// TIA Portal project "SSA-3GHz_V18" (V18) (continued)
REGION Network 4: INFO: If T_CONFIG is done, "start" will be reset.
   RUNG wire#powerrail
      { S7_Templates := "SrcType := DWord" } EQ_Contact(in1 := "SLI_gDB_T_CONFIG_PLC".T_CONFIG.status, in2 := 16#0070_0200)
      R_Coil( "SLI_gDB_T_CONFIG_PLC".T_CONFIG.start )
   END_RUNG
   // the same network as SCL:
   IF "SLI_gDB_T_CONFIG_PLC".T_CONFIG.status = 16#0070_0200 THEN
       "SLI_gDB_T_CONFIG_PLC".T_CONFIG.start := FALSE;
   END_IF;
END_REGION
END_FUNCTION

FUNCTION "ProcessDI" : Void   // FC400, LAD
{ S7_Optimized_Access := 'TRUE' }
VERSION : 0.1
BEGIN

REGION Network 1: DutyCycOK
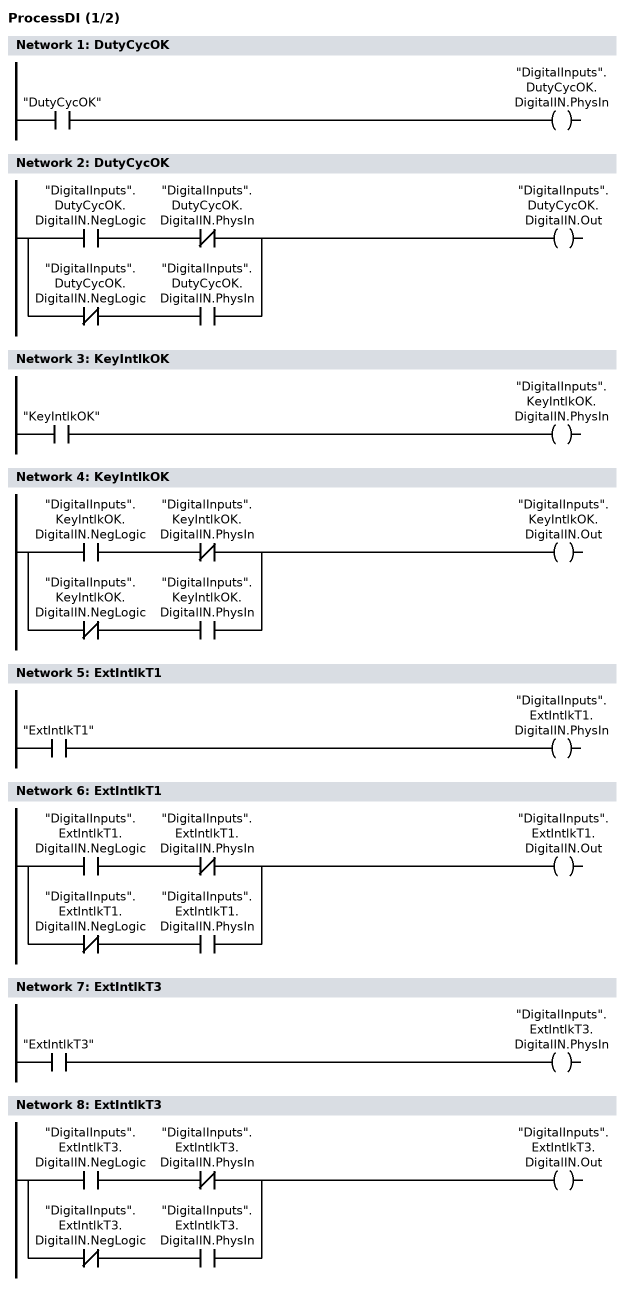
   RUNG wire#powerrail
      Contact( "DutyCycOK" )
      Coil( "DigitalInputs".DutyCycOK.DigitalIN.PhysIn )
   END_RUNG
   // the same network as SCL:
   "DigitalInputs".DutyCycOK.DigitalIN.PhysIn := "DutyCycOK";
END_REGION

REGION Network 2: DutyCycOK
   RUNG wire#powerrail
      Contact( "DigitalInputs".DutyCycOK.DigitalIN.NegLogic )
      I_Contact( "DigitalInputs".DutyCycOK.DigitalIN.PhysIn )
      wire#w1
      Coil( "DigitalInputs".DutyCycOK.DigitalIN.Out )
   END_RUNG
   RUNG wire#powerrail
      I_Contact( "DigitalInputs".DutyCycOK.DigitalIN.NegLogic )
      Contact( "DigitalInputs".DutyCycOK.DigitalIN.PhysIn )
   END_RUNG wire#w1
   // the same network as SCL:
   "DigitalInputs".DutyCycOK.DigitalIN.Out := ("DigitalInputs".DutyCycOK.DigitalIN.NegLogic AND NOT "DigitalInputs".DutyCycOK.DigitalIN.PhysIn) OR (NOT "DigitalInputs".DutyCycOK.DigitalIN.NegLogic AND "DigitalInputs".DutyCycOK.DigitalIN.PhysIn);
END_REGION

REGION Network 3: KeyIntlkOK
   RUNG wire#powerrail
      Contact( "KeyIntlkOK" )
      Coil( "DigitalInputs".KeyIntlkOK.DigitalIN.PhysIn )
   END_RUNG
   // the same network as SCL:
   "DigitalInputs".KeyIntlkOK.DigitalIN.PhysIn := "KeyIntlkOK";
END_REGION

REGION Network 4: KeyIntlkOK
   RUNG wire#powerrail
      Contact( "DigitalInputs".KeyIntlkOK.DigitalIN.NegLogic )
      I_Contact( "DigitalInputs".KeyIntlkOK.DigitalIN.PhysIn )
      wire#w1
      Coil( "DigitalInputs".KeyIntlkOK.DigitalIN.Out )
   END_RUNG
   RUNG wire#powerrail
      I_Contact( "DigitalInputs".KeyIntlkOK.DigitalIN.NegLogic )
      Contact( "DigitalInputs".KeyIntlkOK.DigitalIN.PhysIn )
   END_RUNG wire#w1
   // the same network as SCL:
   "DigitalInputs".KeyIntlkOK.DigitalIN.Out := ("DigitalInputs".KeyIntlkOK.DigitalIN.NegLogic AND NOT "DigitalInputs".KeyIntlkOK.DigitalIN.PhysIn) OR (NOT "DigitalInputs".KeyIntlkOK.DigitalIN.NegLogic AND "DigitalInputs".KeyIntlkOK.DigitalIN.PhysIn);
END_REGION

REGION Network 5: ExtIntlkT1
   RUNG wire#powerrail
      Contact( "ExtIntlkT1" )
      Coil( "DigitalInputs".ExtIntlkT1.DigitalIN.PhysIn )
   END_RUNG
   // the same network as SCL:
   "DigitalInputs".ExtIntlkT1.DigitalIN.PhysIn := "ExtIntlkT1";
END_REGION

REGION Network 6: ExtIntlkT1
   RUNG wire#powerrail
      Contact( "DigitalInputs".ExtIntlkT1.DigitalIN.NegLogic )
      I_Contact( "DigitalInputs".ExtIntlkT1.DigitalIN.PhysIn )
      wire#w1
      Coil( "DigitalInputs".ExtIntlkT1.DigitalIN.Out )
   END_RUNG
   RUNG wire#powerrail
      I_Contact( "DigitalInputs".ExtIntlkT1.DigitalIN.NegLogic )
      Contact( "DigitalInputs".ExtIntlkT1.DigitalIN.PhysIn )
   END_RUNG wire#w1
   // the same network as SCL:
   "DigitalInputs".ExtIntlkT1.DigitalIN.Out := ("DigitalInputs".ExtIntlkT1.DigitalIN.NegLogic AND NOT "DigitalInputs".ExtIntlkT1.DigitalIN.PhysIn) OR (NOT "DigitalInputs".ExtIntlkT1.DigitalIN.NegLogic AND "DigitalInputs".ExtIntlkT1.DigitalIN.PhysIn);
END_REGION

REGION Network 7: ExtIntlkT3
   RUNG wire#powerrail
      Contact( "ExtIntlkT3" )
      Coil( "DigitalInputs".ExtIntlkT3.DigitalIN.PhysIn )
   END_RUNG
   // the same network as SCL:
   "DigitalInputs".ExtIntlkT3.DigitalIN.PhysIn := "ExtIntlkT3";
END_REGION

REGION Network 8: ExtIntlkT3
   RUNG wire#powerrail
      Contact( "DigitalInputs".ExtIntlkT3.DigitalIN.NegLogic )
      I_Contact( "DigitalInputs".ExtIntlkT3.DigitalIN.PhysIn )
      wire#w1
      Coil( "DigitalInputs".ExtIntlkT3.DigitalIN.Out )
   END_RUNG
   RUNG wire#powerrail
      I_Contact( "DigitalInputs".ExtIntlkT3.DigitalIN.NegLogic )
      Contact( "DigitalInputs".ExtIntlkT3.DigitalIN.PhysIn )
   END_RUNG wire#w1
   // the same network as SCL:
   "DigitalInputs".ExtIntlkT3.DigitalIN.Out := ("DigitalInputs".ExtIntlkT3.DigitalIN.NegLogic AND NOT "DigitalInputs".ExtIntlkT3.DigitalIN.PhysIn) OR (NOT "DigitalInputs".ExtIntlkT3.DigitalIN.NegLogic AND "DigitalInputs".ExtIntlkT3.DigitalIN.PhysIn);
END_REGION

REGION Network 9: PS_OK
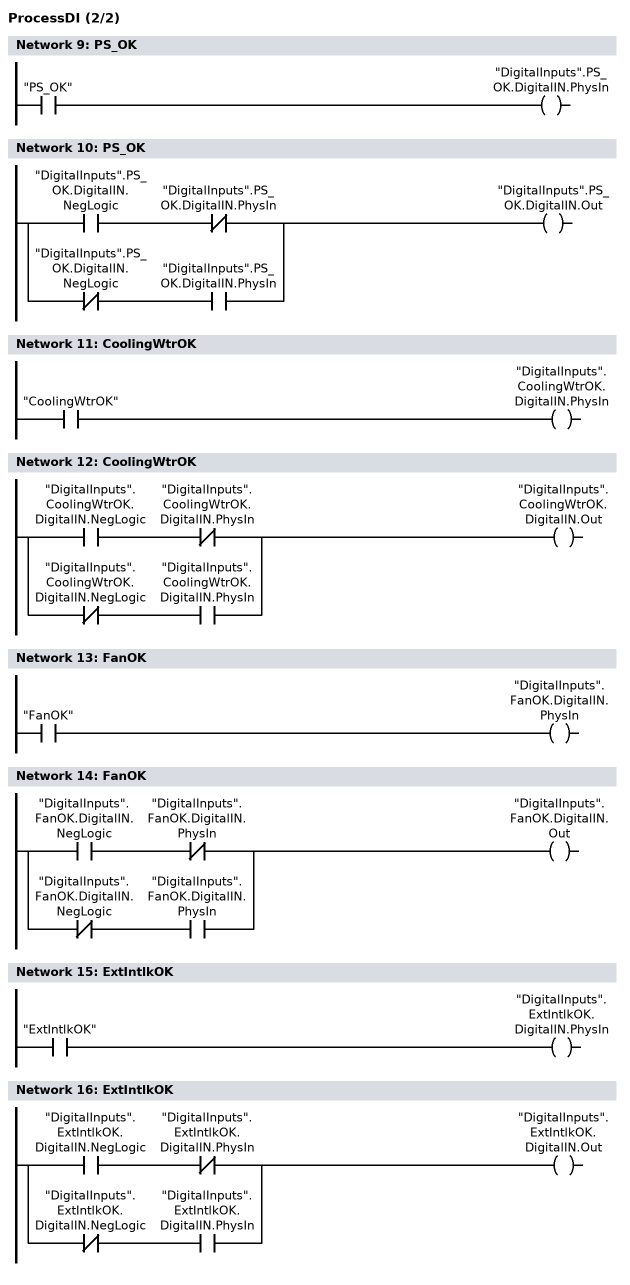
   RUNG wire#powerrail
      Contact( "PS_OK" )
      Coil( "DigitalInputs".PS_OK.DigitalIN.PhysIn )
   END_RUNG
   // the same network as SCL:
   "DigitalInputs".PS_OK.DigitalIN.PhysIn := "PS_OK";
END_REGION

REGION Network 10: PS_OK
   RUNG wire#powerrail
      Contact( "DigitalInputs".PS_OK.DigitalIN.NegLogic )
      I_Contact( "DigitalInputs".PS_OK.DigitalIN.PhysIn )
      wire#w1
      Coil( "DigitalInputs".PS_OK.DigitalIN.Out )
   END_RUNG
   RUNG wire#powerrail
      I_Contact( "DigitalInputs".PS_OK.DigitalIN.NegLogic )
      Contact( "DigitalInputs".PS_OK.DigitalIN.PhysIn )
   END_RUNG wire#w1
   // the same network as SCL:
   "DigitalInputs".PS_OK.DigitalIN.Out := ("DigitalInputs".PS_OK.DigitalIN.NegLogic AND NOT "DigitalInputs".PS_OK.DigitalIN.PhysIn) OR (NOT "DigitalInputs".PS_OK.DigitalIN.NegLogic AND "DigitalInputs".PS_OK.DigitalIN.PhysIn);
END_REGION

REGION Network 11: CoolingWtrOK
   RUNG wire#powerrail
      Contact( "CoolingWtrOK" )
      Coil( "DigitalInputs".CoolingWtrOK.DigitalIN.PhysIn )
   END_RUNG
   // the same network as SCL:
   "DigitalInputs".CoolingWtrOK.DigitalIN.PhysIn := "CoolingWtrOK";
END_REGION

REGION Network 12: CoolingWtrOK
   RUNG wire#powerrail
      Contact( "DigitalInputs".CoolingWtrOK.DigitalIN.NegLogic )
      I_Contact( "DigitalInputs".CoolingWtrOK.DigitalIN.PhysIn )
      wire#w1
      Coil( "DigitalInputs".CoolingWtrOK.DigitalIN.Out )
   END_RUNG
   RUNG wire#powerrail
      I_Contact( "DigitalInputs".CoolingWtrOK.DigitalIN.NegLogic )
      Contact( "DigitalInputs".CoolingWtrOK.DigitalIN.PhysIn )
   END_RUNG wire#w1
   // the same network as SCL:
   "DigitalInputs".CoolingWtrOK.DigitalIN.Out := ("DigitalInputs".CoolingWtrOK.DigitalIN.NegLogic AND NOT "DigitalInputs".CoolingWtrOK.DigitalIN.PhysIn) OR (NOT "DigitalInputs".CoolingWtrOK.DigitalIN.NegLogic AND "DigitalInputs".CoolingWtrOK.DigitalIN.PhysIn);
END_REGION

REGION Network 13: FanOK
   RUNG wire#powerrail
      Contact( "FanOK" )
      Coil( "DigitalInputs".FanOK.DigitalIN.PhysIn )
   END_RUNG
   // the same network as SCL:
   "DigitalInputs".FanOK.DigitalIN.PhysIn := "FanOK";
END_REGION

REGION Network 14: FanOK
   RUNG wire#powerrail
      Contact( "DigitalInputs".FanOK.DigitalIN.NegLogic )
      I_Contact( "DigitalInputs".FanOK.DigitalIN.PhysIn )
      wire#w1
      Coil( "DigitalInputs".FanOK.DigitalIN.Out )
   END_RUNG
   RUNG wire#powerrail
      I_Contact( "DigitalInputs".FanOK.DigitalIN.NegLogic )
      Contact( "DigitalInputs".FanOK.DigitalIN.PhysIn )
   END_RUNG wire#w1
   // the same network as SCL:
   "DigitalInputs".FanOK.DigitalIN.Out := ("DigitalInputs".FanOK.DigitalIN.NegLogic AND NOT "DigitalInputs".FanOK.DigitalIN.PhysIn) OR (NOT "DigitalInputs".FanOK.DigitalIN.NegLogic AND "DigitalInputs".FanOK.DigitalIN.PhysIn);
END_REGION

REGION Network 15: ExtIntlkOK
   RUNG wire#powerrail
      Contact( "ExtIntlkOK" )
      Coil( "DigitalInputs".ExtIntlkOK.DigitalIN.PhysIn )
   END_RUNG
   // the same network as SCL:
   "DigitalInputs".ExtIntlkOK.DigitalIN.PhysIn := "ExtIntlkOK";
END_REGION

REGION Network 16: ExtIntlkOK
   RUNG wire#powerrail
      Contact( "DigitalInputs".ExtIntlkOK.DigitalIN.NegLogic )
      I_Contact( "DigitalInputs".ExtIntlkOK.DigitalIN.PhysIn )
      wire#w1
      Coil( "DigitalInputs".ExtIntlkOK.DigitalIN.Out )
   END_RUNG
   RUNG wire#powerrail
      I_Contact( "DigitalInputs".ExtIntlkOK.DigitalIN.NegLogic )
      Contact( "DigitalInputs".ExtIntlkOK.DigitalIN.PhysIn )
   END_RUNG wire#w1
   // the same network as SCL:
   "DigitalInputs".ExtIntlkOK.DigitalIN.Out := ("DigitalInputs".ExtIntlkOK.DigitalIN.NegLogic AND NOT "DigitalInputs".ExtIntlkOK.DigitalIN.PhysIn) OR (NOT "DigitalInputs".ExtIntlkOK.DigitalIN.NegLogic AND "DigitalInputs".ExtIntlkOK.DigitalIN.PhysIn);
END_REGION
END_FUNCTION

FUNCTION "ProcessAI" : Void   // FC401, LAD
{ S7_Optimized_Access := 'TRUE' }
VERSION : 0.1
   VAR_TEMP
      tmpR1 : Real;
      tmpR : Real;
   END_VAR
BEGIN

REGION Network 1: U drain_RBK
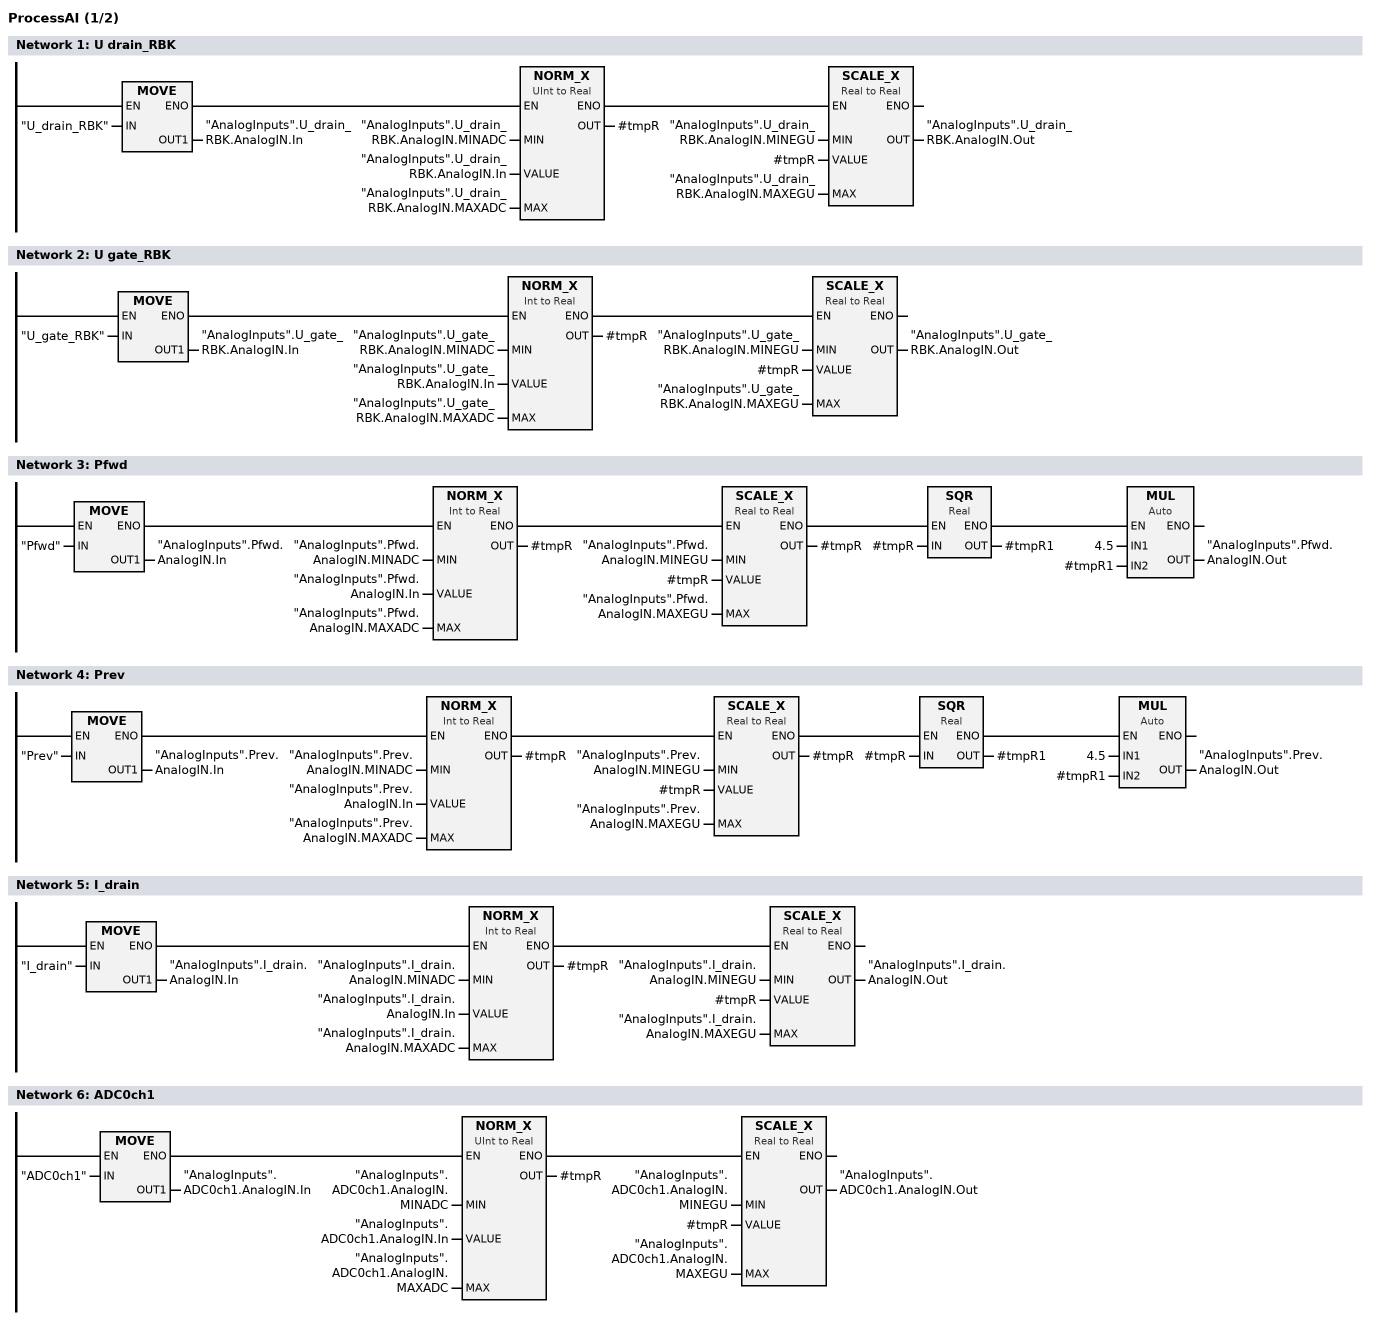
   RUNG wire#powerrail
      Move(in := "U_drain_RBK", out1 => "AnalogInputs".U_drain_RBK.AnalogIN.In)
      { S7_Templates := "[SrcType := UInt, DestType := Real]" } Normalize(min := "AnalogInputs".U_drain_RBK.AnalogIN.MINADC, value := "AnalogInputs".U_drain_RBK.AnalogIN.In, max := "AnalogInputs".U_drain_RBK.AnalogIN.MAXADC, out => #tmpR)
      { S7_Templates := "[SrcType := Real, DestType := Real]" } Scale(min := "AnalogInputs".U_drain_RBK.AnalogIN.MINEGU, value := #tmpR, max := "AnalogInputs".U_drain_RBK.AnalogIN.MAXEGU, out => "AnalogInputs".U_drain_RBK.AnalogIN.Out)
   END_RUNG
   // the same network as SCL:
   "AnalogInputs".U_drain_RBK.AnalogIN.In := "U_drain_RBK";
   #tmpR := NORM_X(MIN := "AnalogInputs".U_drain_RBK.AnalogIN.MINADC, VALUE := "AnalogInputs".U_drain_RBK.AnalogIN.In, MAX := "AnalogInputs".U_drain_RBK.AnalogIN.MAXADC);
   "AnalogInputs".U_drain_RBK.AnalogIN.Out := SCALE_X(MIN := "AnalogInputs".U_drain_RBK.AnalogIN.MINEGU, VALUE := #tmpR, MAX := "AnalogInputs".U_drain_RBK.AnalogIN.MAXEGU);
END_REGION

REGION Network 2: U gate_RBK
   RUNG wire#powerrail
      Move(in := "U_gate_RBK", out1 => "AnalogInputs".U_gate_RBK.AnalogIN.In)
      { S7_Templates := "[SrcType := Int, DestType := Real]" } Normalize(min := "AnalogInputs".U_gate_RBK.AnalogIN.MINADC, value := "AnalogInputs".U_gate_RBK.AnalogIN.In, max := "AnalogInputs".U_gate_RBK.AnalogIN.MAXADC, out => #tmpR)
      { S7_Templates := "[SrcType := Real, DestType := Real]" } Scale(min := "AnalogInputs".U_gate_RBK.AnalogIN.MINEGU, value := #tmpR, max := "AnalogInputs".U_gate_RBK.AnalogIN.MAXEGU, out => "AnalogInputs".U_gate_RBK.AnalogIN.Out)
   END_RUNG
   // the same network as SCL:
   "AnalogInputs".U_gate_RBK.AnalogIN.In := "U_gate_RBK";
   #tmpR := NORM_X(MIN := "AnalogInputs".U_gate_RBK.AnalogIN.MINADC, VALUE := "AnalogInputs".U_gate_RBK.AnalogIN.In, MAX := "AnalogInputs".U_gate_RBK.AnalogIN.MAXADC);
   "AnalogInputs".U_gate_RBK.AnalogIN.Out := SCALE_X(MIN := "AnalogInputs".U_gate_RBK.AnalogIN.MINEGU, VALUE := #tmpR, MAX := "AnalogInputs".U_gate_RBK.AnalogIN.MAXEGU);
END_REGION

REGION Network 3: Pfwd
   "AnalogInputs".Pfwd.AnalogIN.In := "Pfwd";
   #tmpR := NORM_X(MIN := "AnalogInputs".Pfwd.AnalogIN.MINADC, VALUE := "AnalogInputs".Pfwd.AnalogIN.In, MAX := "AnalogInputs".Pfwd.AnalogIN.MAXADC);
   #tmpR := SCALE_X(MIN := "AnalogInputs".Pfwd.AnalogIN.MINEGU, VALUE := #tmpR, MAX := "AnalogInputs".Pfwd.AnalogIN.MAXEGU);
   #tmpR1 := SQR(#tmpR);
   "AnalogInputs".Pfwd.AnalogIN.Out := 4.5 * #tmpR1;
END_REGION

REGION Network 4: Prev
   "AnalogInputs".Prev.AnalogIN.In := "Prev";
   #tmpR := NORM_X(MIN := "AnalogInputs".Prev.AnalogIN.MINADC, VALUE := "AnalogInputs".Prev.AnalogIN.In, MAX := "AnalogInputs".Prev.AnalogIN.MAXADC);
   #tmpR := SCALE_X(MIN := "AnalogInputs".Prev.AnalogIN.MINEGU, VALUE := #tmpR, MAX := "AnalogInputs".Prev.AnalogIN.MAXEGU);
   #tmpR1 := SQR(#tmpR);
   "AnalogInputs".Prev.AnalogIN.Out := 4.5 * #tmpR1;
END_REGION

REGION Network 5: I_drain
   RUNG wire#powerrail
      Move(in := "I_drain", out1 => "AnalogInputs".I_drain.AnalogIN.In)
      { S7_Templates := "[SrcType := Int, DestType := Real]" } Normalize(min := "AnalogInputs".I_drain.AnalogIN.MINADC, value := "AnalogInputs".I_drain.AnalogIN.In, max := "AnalogInputs".I_drain.AnalogIN.MAXADC, out => #tmpR)
      { S7_Templates := "[SrcType := Real, DestType := Real]" } Scale(min := "AnalogInputs".I_drain.AnalogIN.MINEGU, value := #tmpR, max := "AnalogInputs".I_drain.AnalogIN.MAXEGU, out => "AnalogInputs".I_drain.AnalogIN.Out)
   END_RUNG
   // the same network as SCL:
   "AnalogInputs".I_drain.AnalogIN.In := "I_drain";
   #tmpR := NORM_X(MIN := "AnalogInputs".I_drain.AnalogIN.MINADC, VALUE := "AnalogInputs".I_drain.AnalogIN.In, MAX := "AnalogInputs".I_drain.AnalogIN.MAXADC);
   "AnalogInputs".I_drain.AnalogIN.Out := SCALE_X(MIN := "AnalogInputs".I_drain.AnalogIN.MINEGU, VALUE := #tmpR, MAX := "AnalogInputs".I_drain.AnalogIN.MAXEGU);
END_REGION

REGION Network 6: ADC0ch1
   RUNG wire#powerrail
      Move(in := "ADC0ch1", out1 => "AnalogInputs".ADC0ch1.AnalogIN.In)
      { S7_Templates := "[SrcType := UInt, DestType := Real]" } Normalize(min := "AnalogInputs".ADC0ch1.AnalogIN.MINADC, value := "AnalogInputs".ADC0ch1.AnalogIN.In, max := "AnalogInputs".ADC0ch1.AnalogIN.MAXADC, out => #tmpR)
      { S7_Templates := "[SrcType := Real, DestType := Real]" } Scale(min := "AnalogInputs".ADC0ch1.AnalogIN.MINEGU, value := #tmpR, max := "AnalogInputs".ADC0ch1.AnalogIN.MAXEGU, out => "AnalogInputs".ADC0ch1.AnalogIN.Out)
   END_RUNG
   // the same network as SCL:
   "AnalogInputs".ADC0ch1.AnalogIN.In := "ADC0ch1";
   #tmpR := NORM_X(MIN := "AnalogInputs".ADC0ch1.AnalogIN.MINADC, VALUE := "AnalogInputs".ADC0ch1.AnalogIN.In, MAX := "AnalogInputs".ADC0ch1.AnalogIN.MAXADC);
   "AnalogInputs".ADC0ch1.AnalogIN.Out := SCALE_X(MIN := "AnalogInputs".ADC0ch1.AnalogIN.MINEGU, VALUE := #tmpR, MAX := "AnalogInputs".ADC0ch1.AnalogIN.MAXEGU);
END_REGION

REGION Network 7: Pfwd in dBm
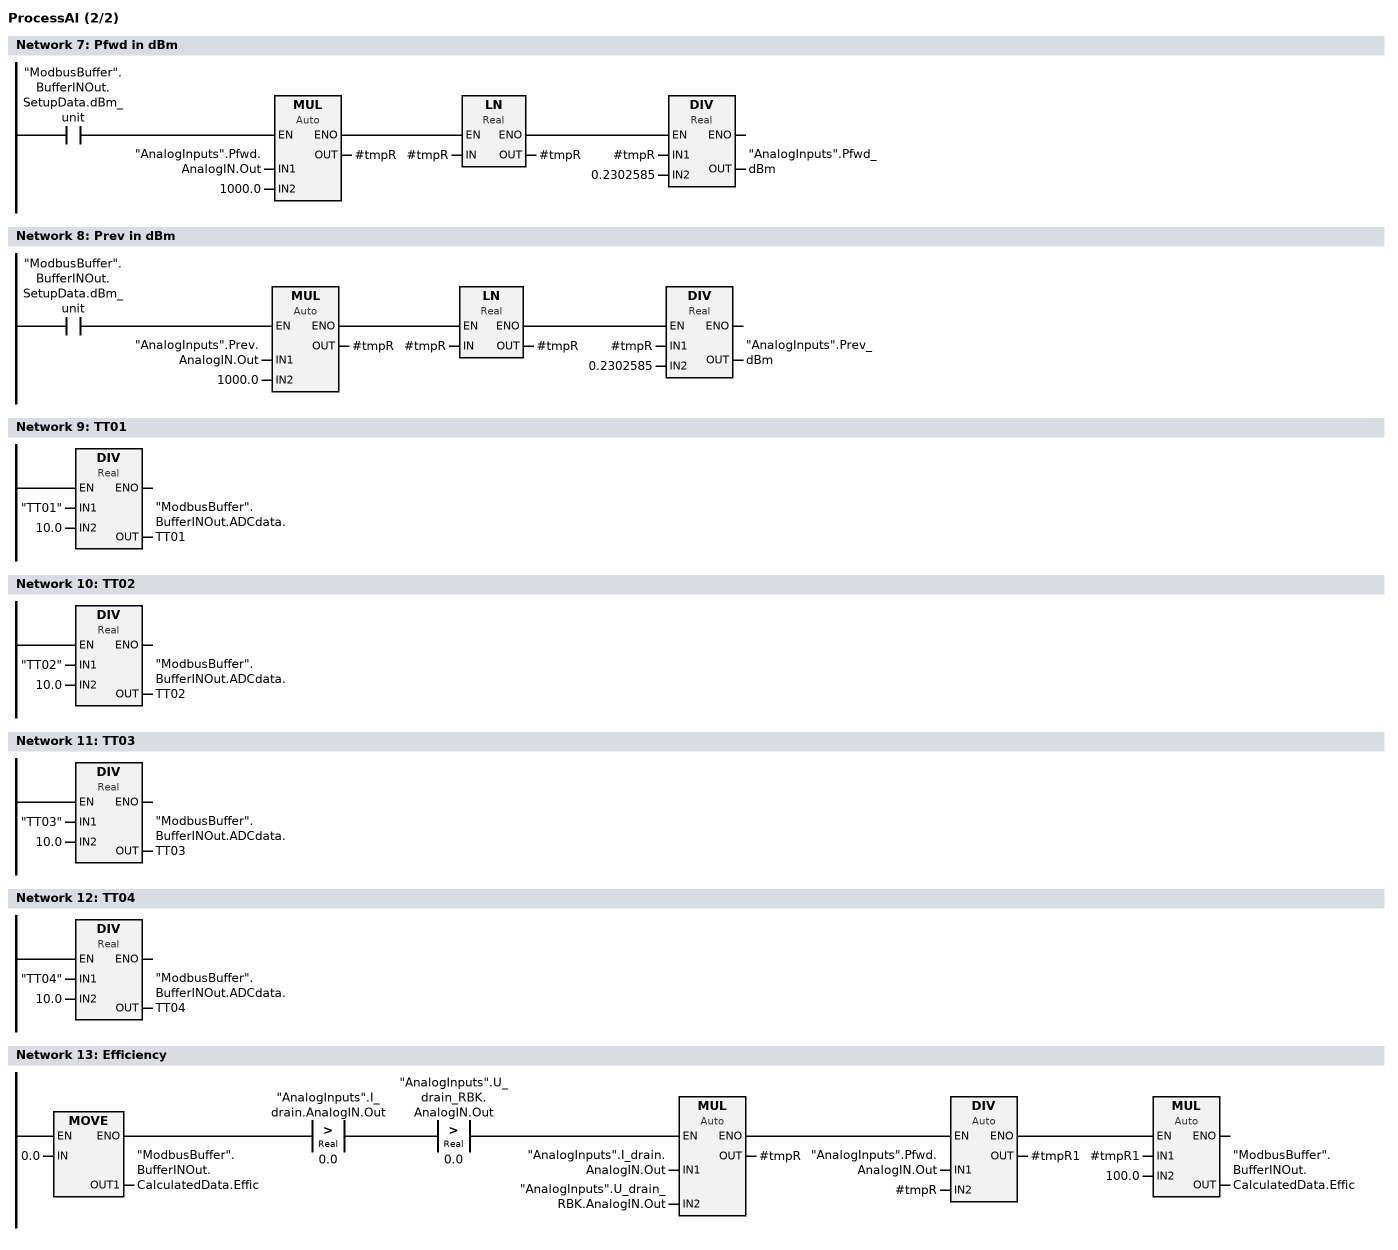
   IF "ModbusBuffer".BufferINOut.SetupData.dBm_unit THEN
       #tmpR := "AnalogInputs".Pfwd.AnalogIN.Out * 1000.0;
       #tmpR := LN(#tmpR);
       "AnalogInputs".Pfwd_dBm := #tmpR / 0.2302585;
   END_IF;
END_REGION

REGION Network 8: Prev in dBm
   IF "ModbusBuffer".BufferINOut.SetupData.dBm_unit THEN
       #tmpR := "AnalogInputs".Prev.AnalogIN.Out * 1000.0;
       #tmpR := LN(#tmpR);
       "AnalogInputs".Prev_dBm := #tmpR / 0.2302585;
   END_IF;
END_REGION

REGION Network 9: TT01
   RUNG wire#powerrail
      { S7_Templates := "SrcType := Real" } Div(in1 := "TT01", in2 := 10.0, out => "ModbusBuffer".BufferINOut.ADCdata.TT01)
   END_RUNG
   // the same network as SCL:
   "ModbusBuffer".BufferINOut.ADCdata.TT01 := "TT01" / 10.0;
END_REGION

REGION Network 10: TT02
   RUNG wire#powerrail
      { S7_Templates := "SrcType := Real" } Div(in1 := "TT02", in2 := 10.0, out => "ModbusBuffer".BufferINOut.ADCdata.TT02)
   END_RUNG
   // the same network as SCL:
   "ModbusBuffer".BufferINOut.ADCdata.TT02 := "TT02" / 10.0;
END_REGION

REGION Network 11: TT03
   RUNG wire#powerrail
      { S7_Templates := "SrcType := Real" } Div(in1 := "TT03", in2 := 10.0, out => "ModbusBuffer".BufferINOut.ADCdata.TT03)
   END_RUNG
   // the same network as SCL:
   "ModbusBuffer".BufferINOut.ADCdata.TT03 := "TT03" / 10.0;
END_REGION

REGION Network 12: TT04
   RUNG wire#powerrail
      { S7_Templates := "SrcType := Real" } Div(in1 := "TT04", in2 := 10.0, out => "ModbusBuffer".BufferINOut.ADCdata.TT04)
   END_RUNG
   // the same network as SCL:
   "ModbusBuffer".BufferINOut.ADCdata.TT04 := "TT04" / 10.0;
END_REGION

REGION Network 13: Efficiency
   RUNG wire#powerrail
      Move(in := 0.0, out1 => "ModbusBuffer".BufferINOut.CalculatedData.Effic)
      { S7_Templates := "SrcType := Real" } GT_Contact(in1 := "AnalogInputs".I_drain.AnalogIN.Out, in2 := 0.0)
      { S7_Templates := "SrcType := Real" } GT_Contact(in1 := "AnalogInputs".U_drain_RBK.AnalogIN.Out, in2 := 0.0)
      Mul(in1 := "AnalogInputs".I_drain.AnalogIN.Out, in2 := "AnalogInputs".U_drain_RBK.AnalogIN.Out, out => #tmpR)
      Div(in1 := "AnalogInputs".Pfwd.AnalogIN.Out, in2 := #tmpR, out => #tmpR1)
      Mul(in1 := #tmpR1, in2 := 100.0, out => "ModbusBuffer".BufferINOut.CalculatedData.Effic)
   END_RUNG
   // the same network as SCL:
   "ModbusBuffer".BufferINOut.CalculatedData.Effic := 0.0;
   IF ("AnalogInputs".I_drain.AnalogIN.Out > 0.0) AND ("AnalogInputs".U_drain_RBK.AnalogIN.Out > 0.0) THEN
       #tmpR := "AnalogInputs".I_drain.AnalogIN.Out * "AnalogInputs".U_drain_RBK.AnalogIN.Out;
       #tmpR1 := "AnalogInputs".Pfwd.AnalogIN.Out / #tmpR;
       "ModbusBuffer".BufferINOut.CalculatedData.Effic := #tmpR1 * 100.0;
   END_IF;
END_REGION
END_FUNCTION

FUNCTION "ProcessAO" : Void   // FC402, LAD
{ S7_Optimized_Access := 'TRUE' }
VERSION : 0.1
   VAR_TEMP
      tmpR : Real;
   END_VAR
BEGIN

REGION Network 1: U drain
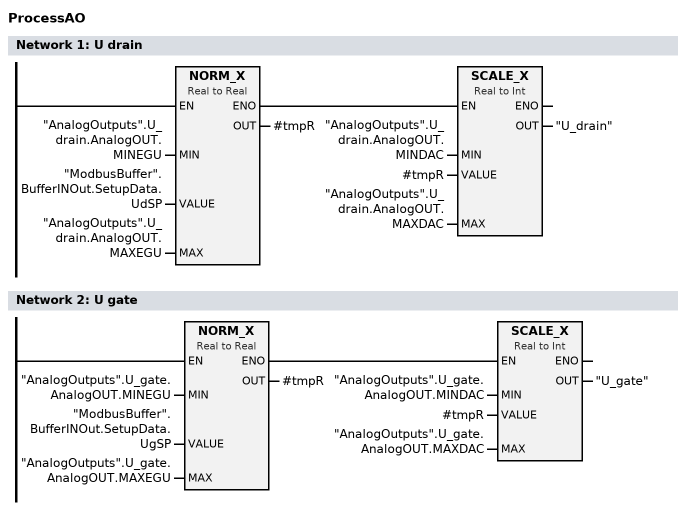
   RUNG wire#powerrail
      { S7_Templates := "[SrcType := Real, DestType := Real]" } Normalize(min := "AnalogOutputs".U_drain.AnalogOUT.MINEGU, value := "ModbusBuffer".BufferINOut.SetupData.UdSP, max := "AnalogOutputs".U_drain.AnalogOUT.MAXEGU, out => #tmpR)
      { S7_Templates := "[SrcType := Real, DestType := Int]" } Scale(min := "AnalogOutputs".U_drain.AnalogOUT.MINDAC, value := #tmpR, max := "AnalogOutputs".U_drain.AnalogOUT.MAXDAC, out => "U_drain")
   END_RUNG
   // the same network as SCL:
   #tmpR := NORM_X(MIN := "AnalogOutputs".U_drain.AnalogOUT.MINEGU, VALUE := "ModbusBuffer".BufferINOut.SetupData.UdSP, MAX := "AnalogOutputs".U_drain.AnalogOUT.MAXEGU);
   "U_drain" := SCALE_X(MIN := "AnalogOutputs".U_drain.AnalogOUT.MINDAC, VALUE := #tmpR, MAX := "AnalogOutputs".U_drain.AnalogOUT.MAXDAC);
END_REGION

REGION Network 2: U gate
   RUNG wire#powerrail
      { S7_Templates := "[SrcType := Real, DestType := Real]" } Normalize(min := "AnalogOutputs".U_gate.AnalogOUT.MINEGU, value := "ModbusBuffer".BufferINOut.SetupData.UgSP, max := "AnalogOutputs".U_gate.AnalogOUT.MAXEGU, out => #tmpR)
      { S7_Templates := "[SrcType := Real, DestType := Int]" } Scale(min := "AnalogOutputs".U_gate.AnalogOUT.MINDAC, value := #tmpR, max := "AnalogOutputs".U_gate.AnalogOUT.MAXDAC, out => "U_gate")
   END_RUNG
   // the same network as SCL:
   #tmpR := NORM_X(MIN := "AnalogOutputs".U_gate.AnalogOUT.MINEGU, VALUE := "ModbusBuffer".BufferINOut.SetupData.UgSP, MAX := "AnalogOutputs".U_gate.AnalogOUT.MAXEGU);
   "U_gate" := SCALE_X(MIN := "AnalogOutputs".U_gate.AnalogOUT.MINDAC, VALUE := #tmpR, MAX := "AnalogOutputs".U_gate.AnalogOUT.MAXDAC);
END_REGION
END_FUNCTION

FUNCTION "ProcessDO" : Void   // FC450, LAD
{ S7_Optimized_Access := 'TRUE' }
VERSION : 0.1
BEGIN

REGION Network 1: RF switcch
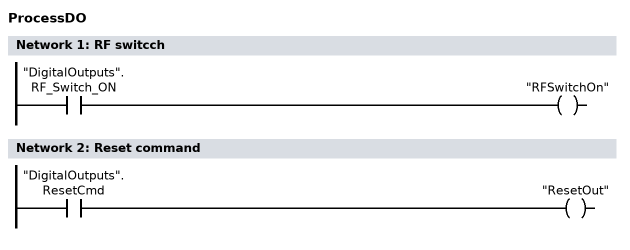
   RUNG wire#powerrail
      Contact( "DigitalOutputs".RF_Switch_ON )
      Coil( "RFSwitchOn" )
   END_RUNG
   // the same network as SCL:
   "RFSwitchOn" := "DigitalOutputs".RF_Switch_ON;
END_REGION

REGION Network 2: Reset command
   RUNG wire#powerrail
      Contact( "DigitalOutputs".ResetCmd )
      Coil( "ResetOut" )
   END_RUNG
   // the same network as SCL:
   "ResetOut" := "DigitalOutputs".ResetCmd;
END_REGION
END_FUNCTION

FUNCTION "CalcTransistorV" : Void   // FC500, SCL
{ S7_Optimized_Access := 'TRUE' }
VERSION : 0.1
   VAR_INPUT
      NominalPwr : Real;
      size : Int;   // max size if the lookup table. Valid data until Pwr != 0
   END_VAR
   VAR_OUTPUT
      UdSP : Real;
      UgSP : Real;
   END_VAR
   VAR_TEMP
      Pwr : Real;
      Ud : Real;
      Ug : Real;
      K : Real;
      i : Int;
   END_VAR
BEGIN
   (*
   Calculate the Darin and gate voltages based on the nominal power
   *)
   IF "ModbusBuffer".BufferINOut.SetupData.dBm_unit THEN
       "ModbusBuffer".BufferINOut.SetupData.NominalPower := EXP("ModbusBuffer".BufferINOut.SetupData.NominalPower_dBm* 0.2302585) / 1000.0;
   ELSE
       "ModbusBuffer".BufferINOut.SetupData.NominalPower_dBm := 10.0 * LN(1000.0 *"ModbusBuffer".BufferINOut.SetupData.NominalPower)/ 2.302585;
   END_IF;

   IF #NominalPwr <= "ModbusBuffer".BufferINOut.LookupTable.Pwr[0] THEN
       #UdSP := "ModbusBuffer".BufferINOut.LookupTable.Ud[0];
       #UgSP := "ModbusBuffer".BufferINOut.LookupTable.Ug[0];
   ELSE
       FOR #i := 1 TO #size-1 DO
       // Statement section FOR
           #Pwr := "ModbusBuffer".BufferINOut.LookupTable.Pwr[#i];
           IF #Pwr = 0 THEN
               //the end of table marker
               #UdSP := "ModbusBuffer".BufferINOut.LookupTable.Ud[#i - 1];
               #UgSP := "ModbusBuffer".BufferINOut.LookupTable.Ug[#i - 1];
               RETURN;
           END_IF;
           IF #NominalPwr > #Pwr THEN
               CONTINUE;
           END_IF;
           #K := (#NominalPwr - "ModbusBuffer".BufferINOut.LookupTable.Pwr[#i - 1]) / (#Pwr - "ModbusBuffer".BufferINOut.LookupTable.Pwr[#i - 1]);
           #UdSP := "ModbusBuffer".BufferINOut.LookupTable.Ud[#i-1] + #K * ("ModbusBuffer".BufferINOut.LookupTable.Ud[#i] - "ModbusBuffer".BufferINOut.LookupTable.Ud[#i-1]);
           #UgSP := "ModbusBuffer".BufferINOut.LookupTable.Ug[#i - 1] + #K * ("ModbusBuffer".BufferINOut.LookupTable.Ug[#i] - "ModbusBuffer".BufferINOut.LookupTable.Ug[#i - 1]);
           RETURN;
       END_FOR;
       #UdSP := "ModbusBuffer".BufferINOut.LookupTable.Ud[#size-1];
       #UgSP := "ModbusBuffer".BufferINOut.LookupTable.Ug[#size-1];
   END_IF;
END_FUNCTION

FUNCTION "Interlocks" : Void   // FC600, LAD
{ S7_Optimized_Access := 'TRUE' }
VERSION : 0.1
BEGIN

REGION Network 1: RF Switch